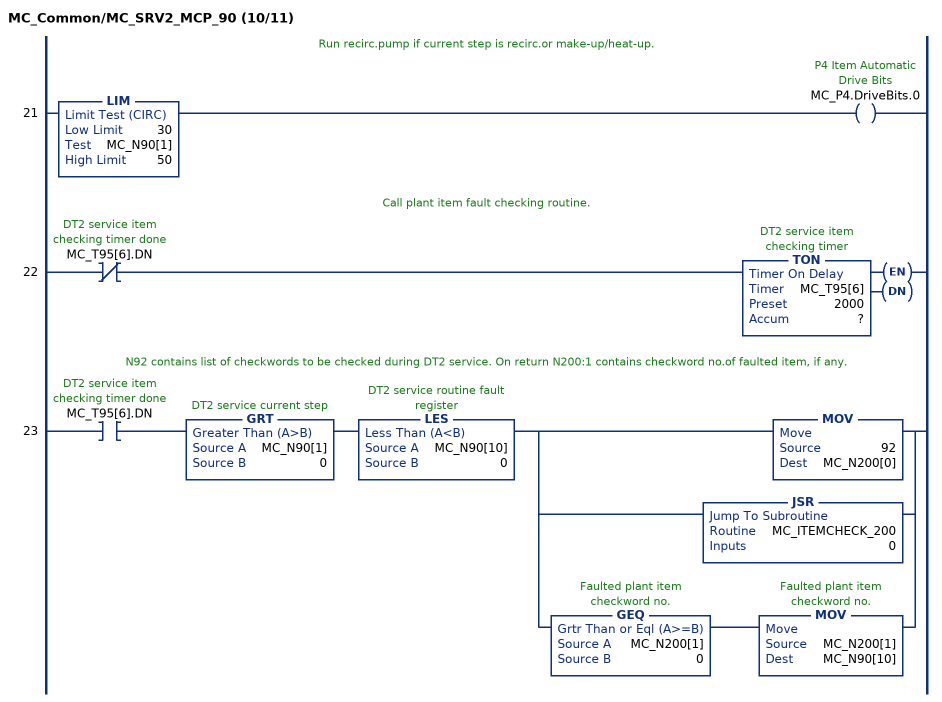
   // Run recirc.pump if current step is recirc.or make-up/heat-up.
   21: LIM(30,MC_N90[1],50)OTE(MC_P4.DriveBits.0);
   // Call plant item fault checking routine.
   22: XIO(MC_T95[6].DN)TON(MC_T95[6],?,?);
   // N92 contains list of checkwords to be checked during DT2 service. On return N200:1 contains checkword no.of faulted item, if any.
   23: XIC(MC_T95[6].DN)GRT(MC_N90[1],0)LES(MC_N90[10],0)[MOV(92,MC_N200[0]) ,JSR(MC_ITEMCHECK_200,0) ,GEQ(MC_N200[1],0) MOV(MC_N200[1],MC_N90[10]) ];
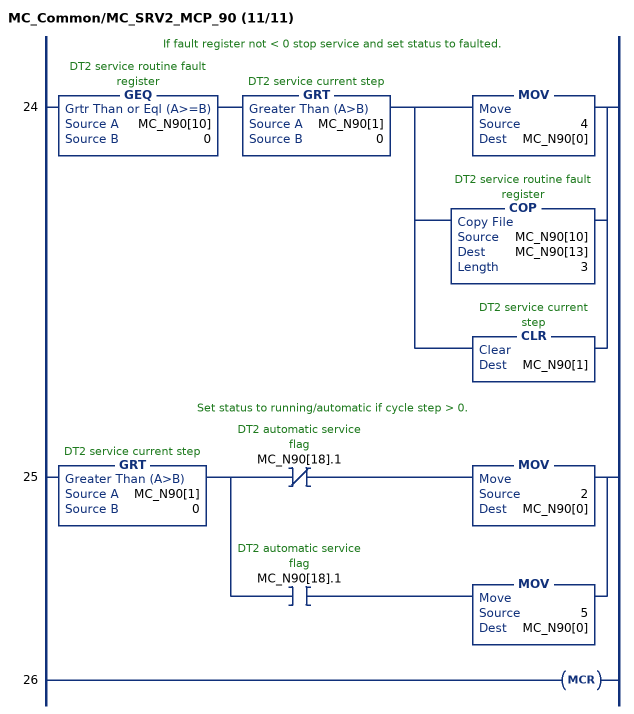
   // If fault register not < 0 stop service and set status to faulted.
   24: GEQ(MC_N90[10],0)GRT(MC_N90[1],0)[MOV(4,MC_N90[0]) ,COP(MC_N90[10],MC_N90[13],3) ,CLR(MC_N90[1]) ];
   // Set status to running/automatic if cycle step > 0.
   25: GRT(MC_N90[1],0)[XIO(MC_N90[18].1) MOV(2,MC_N90[0]) ,XIC(MC_N90[18].1) MOV(5,MC_N90[0]) ];
   26: MCR();
END_ROUTINE

ROUTINE MC_Valves   (* ladder *)
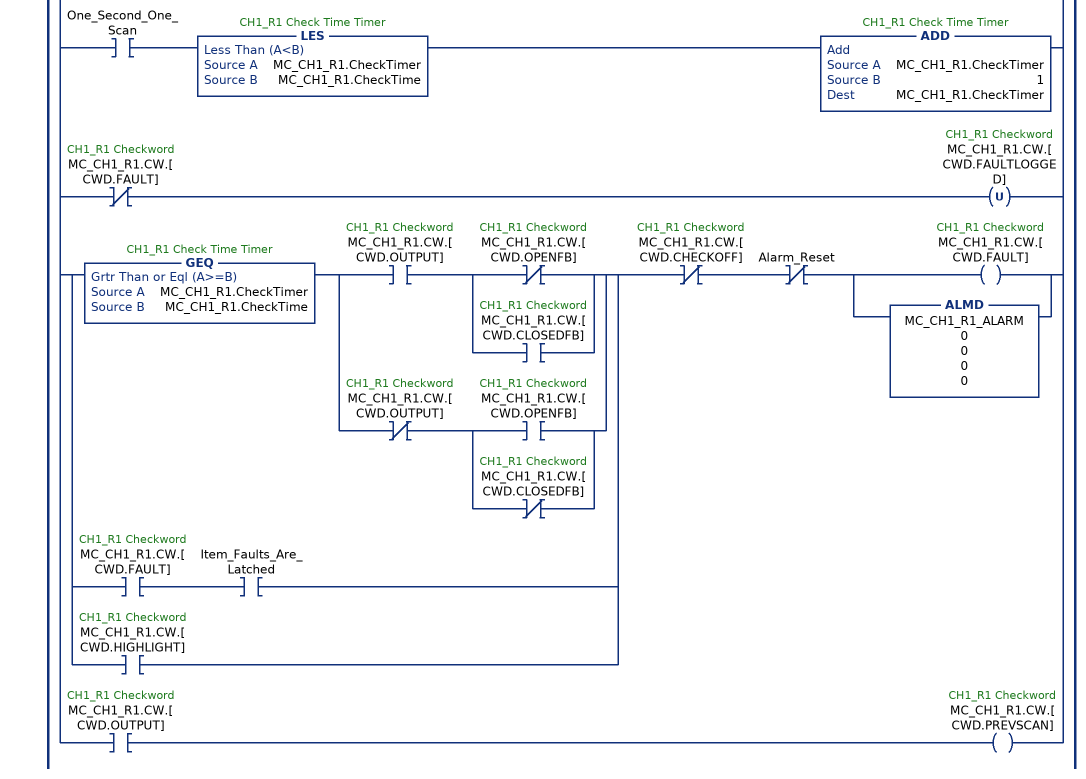
   0: [NEQ(MC_CH1_R1.DriveBits,0) OTE(MC_CH1_R1.CW.[CWD.AUTODRV]) ,[XIC(MC_CH1_R1.CW.[CWD.AUTODRV]) XIO(MC_CH1_R1.CW.[CWD.MANUAL]) ,XIC(MC_CH1_R1.CW.[CWD.MANDRV]) XIC(MC_CH1_R1.CW.[CWD.MANUAL]) ] OTE(MC_CH1_R1.CW.[CWD.OUTPUT]) ,XIC(MC_CH1_R1.CW.[CWD.OUTPUT]) OTE(MC_CH1_R1_DR) ,XIC(S:FS) [OTU(MC_CH1_R1.CW.[CWD.MANUAL]) ,LEQ(MC_CH1_R1.CheckTime,0) MOV(Default_Check_Time,MC_CH1_R1.CheckTime) ] ,[[XIC(MC_CH1_R1_O) XIO(Item_Simulation_Flag) ,XIC(Item_Simulation_Flag) XIC(MC_CH1_R1.CW.[CWD.OUTPUT]) XIO(MC_CH1_R1.CW.[CWD.SIMFAIL]) ] OTE(MC_CH1_R1.CW.[CWD.OPENFB]) ,[XIC(MC_CH1_R1_C) XIO(Item_Simulation_Flag) ,XIC(Item_Simulation_Flag) XIO(MC_CH1_R1.CW.[CWD.OUTPUT]) XIO(MC_CH1_R1.CW.[CWD.SIMFAIL]) ] OTE(MC_CH1_R1.CW.[CWD.CLOSEDFB]) ] ,[XIC(MC_CH1_R1.CW.[CWD.OUTPUT]) XIO(MC_CH1_R1.CW.[CWD.PREVSCAN]) ,XIO(MC_CH1_R1.CW.[CWD.OUTPUT]) XIC(MC_CH1_R1.CW.[CWD.PREVSCAN]) ] CLR(MC_CH1_R1.CheckTimer) ,XIC(One_Second_One_Scan) LES(MC_CH1_R1.CheckTimer,MC_CH1_R1.CheckTime) ADD(MC_CH1_R1.CheckTimer,1,MC_CH1_R1.CheckTimer) ,XIO(MC_CH1_R1.CW.[CWD.FAULT]) OTU(MC_CH1_R1.CW.[CWD.FAULTLOGGED]) ,[GEQ(MC_CH1_R1.CheckTimer,MC_CH1_R1.CheckTime) [XIC(MC_CH1_R1.CW.[CWD.OUTPUT]) [XIO(MC_CH1_R1.CW.[CWD.OPENFB]) ,XIC(MC_CH1_R1.CW.[CWD.CLOSEDFB]) ] ,XIO(MC_CH1_R1.CW.[CWD.OUTPUT]) [XIC(MC_CH1_R1.CW.[CWD.OPENFB]) ,XIO(MC_CH1_R1.CW.[CWD.CLOSEDFB]) ] ] ,XIC(MC_CH1_R1.CW.[CWD.FAULT]) XIC(Item_Faults_Are_Latched) ,XIC(MC_CH1_R1.CW.[CWD.HIGHLIGHT]) ] XIO(MC_CH1_R1.CW.[CWD.CHECKOFF]) XIO(Alarm_Reset) [OTE(MC_CH1_R1.CW.[CWD.FAULT]) ,ALMD(MC_CH1_R1_ALARM,0,0,0,0) ] ,XIC(MC_CH1_R1.CW.[CWD.OUTPUT]) OTE(MC_CH1_R1.CW.[CWD.PREVSCAN]) ];
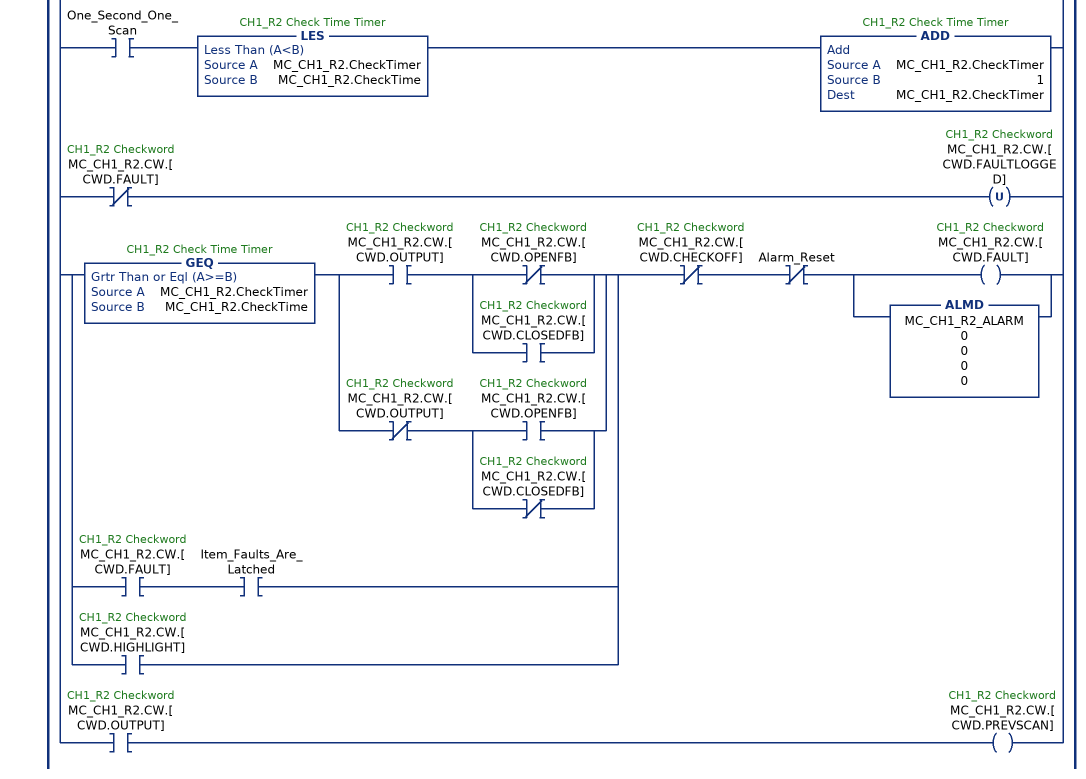
   1: [NEQ(MC_CH1_R2.DriveBits,0) OTE(MC_CH1_R2.CW.[CWD.AUTODRV]) ,[XIC(MC_CH1_R2.CW.[CWD.AUTODRV]) XIO(MC_CH1_R2.CW.[CWD.MANUAL]) ,XIC(MC_CH1_R2.CW.[CWD.MANDRV]) XIC(MC_CH1_R2.CW.[CWD.MANUAL]) ] OTE(MC_CH1_R2.CW.[CWD.OUTPUT]) ,XIC(MC_CH1_R2.CW.[CWD.OUTPUT]) OTE(MC_CH1_R2_DR) ,XIC(S:FS) [OTU(MC_CH1_R2.CW.[CWD.MANUAL]) ,LEQ(MC_CH1_R2.CheckTime,0) MOV(Default_Check_Time,MC_CH1_R2.CheckTime) ] ,[[XIC(MC_CH1_R2_O) XIO(Item_Simulation_Flag) ,XIC(Item_Simulation_Flag) XIC(MC_CH1_R2.CW.[CWD.OUTPUT]) XIO(MC_CH1_R2.CW.[CWD.SIMFAIL]) ] OTE(MC_CH1_R2.CW.[CWD.OPENFB]) ,[XIC(MC_CH1_R2_C) XIO(Item_Simulation_Flag) ,XIC(Item_Simulation_Flag) XIO(MC_CH1_R2.CW.[CWD.OUTPUT]) XIO(MC_CH1_R2.CW.[CWD.SIMFAIL]) ] OTE(MC_CH1_R2.CW.[CWD.CLOSEDFB]) ] ,[XIC(MC_CH1_R2.CW.[CWD.OUTPUT]) XIO(MC_CH1_R2.CW.[CWD.PREVSCAN]) ,XIO(MC_CH1_R2.CW.[CWD.OUTPUT]) XIC(MC_CH1_R2.CW.[CWD.PREVSCAN]) ] CLR(MC_CH1_R2.CheckTimer) ,XIC(One_Second_One_Scan) LES(MC_CH1_R2.CheckTimer,MC_CH1_R2.CheckTime) ADD(MC_CH1_R2.CheckTimer,1,MC_CH1_R2.CheckTimer) ,XIO(MC_CH1_R2.CW.[CWD.FAULT]) OTU(MC_CH1_R2.CW.[CWD.FAULTLOGGED]) ,[GEQ(MC_CH1_R2.CheckTimer,MC_CH1_R2.CheckTime) [XIC(MC_CH1_R2.CW.[CWD.OUTPUT]) [XIO(MC_CH1_R2.CW.[CWD.OPENFB]) ,XIC(MC_CH1_R2.CW.[CWD.CLOSEDFB]) ] ,XIO(MC_CH1_R2.CW.[CWD.OUTPUT]) [XIC(MC_CH1_R2.CW.[CWD.OPENFB]) ,XIO(MC_CH1_R2.CW.[CWD.CLOSEDFB]) ] ] ,XIC(MC_CH1_R2.CW.[CWD.FAULT]) XIC(Item_Faults_Are_Latched) ,XIC(MC_CH1_R2.CW.[CWD.HIGHLIGHT]) ] XIO(MC_CH1_R2.CW.[CWD.CHECKOFF]) XIO(Alarm_Reset) [OTE(MC_CH1_R2.CW.[CWD.FAULT]) ,ALMD(MC_CH1_R2_ALARM,0,0,0,0) ] ,XIC(MC_CH1_R2.CW.[CWD.OUTPUT]) OTE(MC_CH1_R2.CW.[CWD.PREVSCAN]) ];
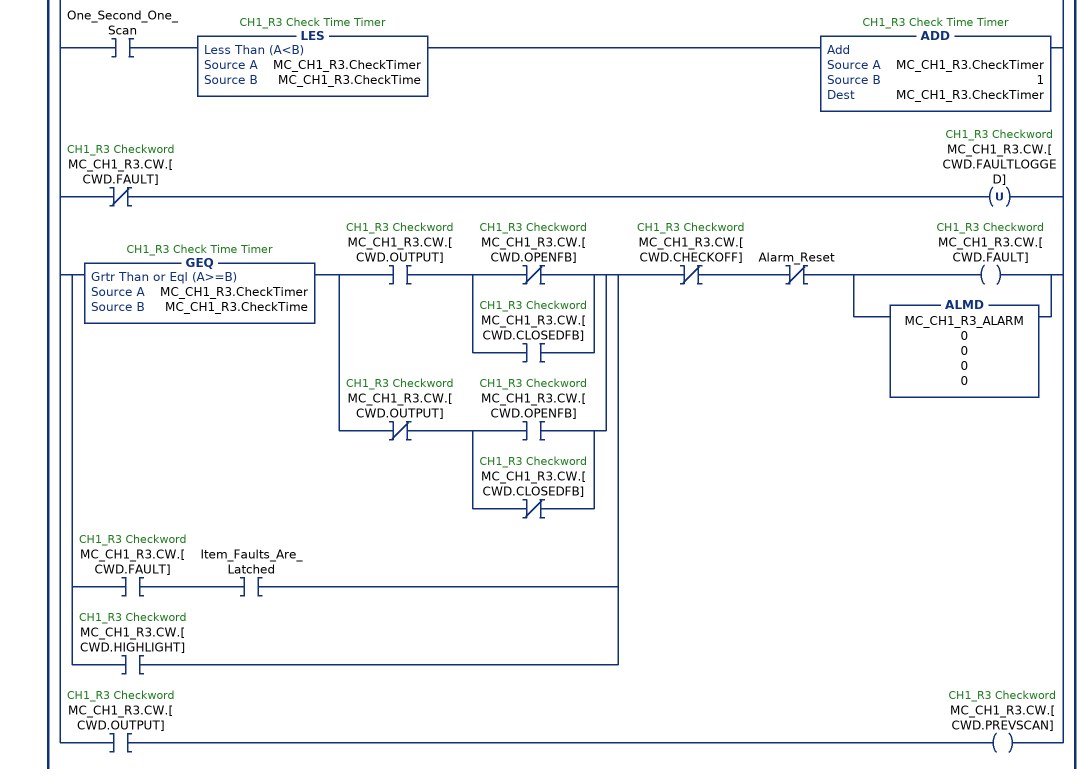
   2: [NEQ(MC_CH1_R3.DriveBits,0) OTE(MC_CH1_R3.CW.[CWD.AUTODRV]) ,[XIC(MC_CH1_R3.CW.[CWD.AUTODRV]) XIO(MC_CH1_R3.CW.[CWD.MANUAL]) ,XIC(MC_CH1_R3.CW.[CWD.MANDRV]) XIC(MC_CH1_R3.CW.[CWD.MANUAL]) ] OTE(MC_CH1_R3.CW.[CWD.OUTPUT]) ,XIC(MC_CH1_R3.CW.[CWD.OUTPUT]) OTE(MC_CH1_R3_DR) ,XIC(S:FS) [OTU(MC_CH1_R3.CW.[CWD.MANUAL]) ,LEQ(MC_CH1_R3.CheckTime,0) MOV(Default_Check_Time,MC_CH1_R3.CheckTime) ] ,[[XIC(MC_CH1_R3_O) XIO(Item_Simulation_Flag) ,XIC(Item_Simulation_Flag) XIC(MC_CH1_R3.CW.[CWD.OUTPUT]) XIO(MC_CH1_R3.CW.[CWD.SIMFAIL]) ] OTE(MC_CH1_R3.CW.[CWD.OPENFB]) ,[XIC(MC_CH1_R3_C) XIO(Item_Simulation_Flag) ,XIC(Item_Simulation_Flag) XIO(MC_CH1_R3.CW.[CWD.OUTPUT]) XIO(MC_CH1_R3.CW.[CWD.SIMFAIL]) ] OTE(MC_CH1_R3.CW.[CWD.CLOSEDFB]) ] ,[XIC(MC_CH1_R3.CW.[CWD.OUTPUT]) XIO(MC_CH1_R3.CW.[CWD.PREVSCAN]) ,XIO(MC_CH1_R3.CW.[CWD.OUTPUT]) XIC(MC_CH1_R3.CW.[CWD.PREVSCAN]) ] CLR(MC_CH1_R3.CheckTimer) ,XIC(One_Second_One_Scan) LES(MC_CH1_R3.CheckTimer,MC_CH1_R3.CheckTime) ADD(MC_CH1_R3.CheckTimer,1,MC_CH1_R3.CheckTimer) ,XIO(MC_CH1_R3.CW.[CWD.FAULT]) OTU(MC_CH1_R3.CW.[CWD.FAULTLOGGED]) ,[GEQ(MC_CH1_R3.CheckTimer,MC_CH1_R3.CheckTime) [XIC(MC_CH1_R3.CW.[CWD.OUTPUT]) [XIO(MC_CH1_R3.CW.[CWD.OPENFB]) ,XIC(MC_CH1_R3.CW.[CWD.CLOSEDFB]) ] ,XIO(MC_CH1_R3.CW.[CWD.OUTPUT]) [XIC(MC_CH1_R3.CW.[CWD.OPENFB]) ,XIO(MC_CH1_R3.CW.[CWD.CLOSEDFB]) ] ] ,XIC(MC_CH1_R3.CW.[CWD.FAULT]) XIC(Item_Faults_Are_Latched) ,XIC(MC_CH1_R3.CW.[CWD.HIGHLIGHT]) ] XIO(MC_CH1_R3.CW.[CWD.CHECKOFF]) XIO(Alarm_Reset) [OTE(MC_CH1_R3.CW.[CWD.FAULT]) ,ALMD(MC_CH1_R3_ALARM,0,0,0,0) ] ,XIC(MC_CH1_R3.CW.[CWD.OUTPUT]) OTE(MC_CH1_R3.CW.[CWD.PREVSCAN]) ];
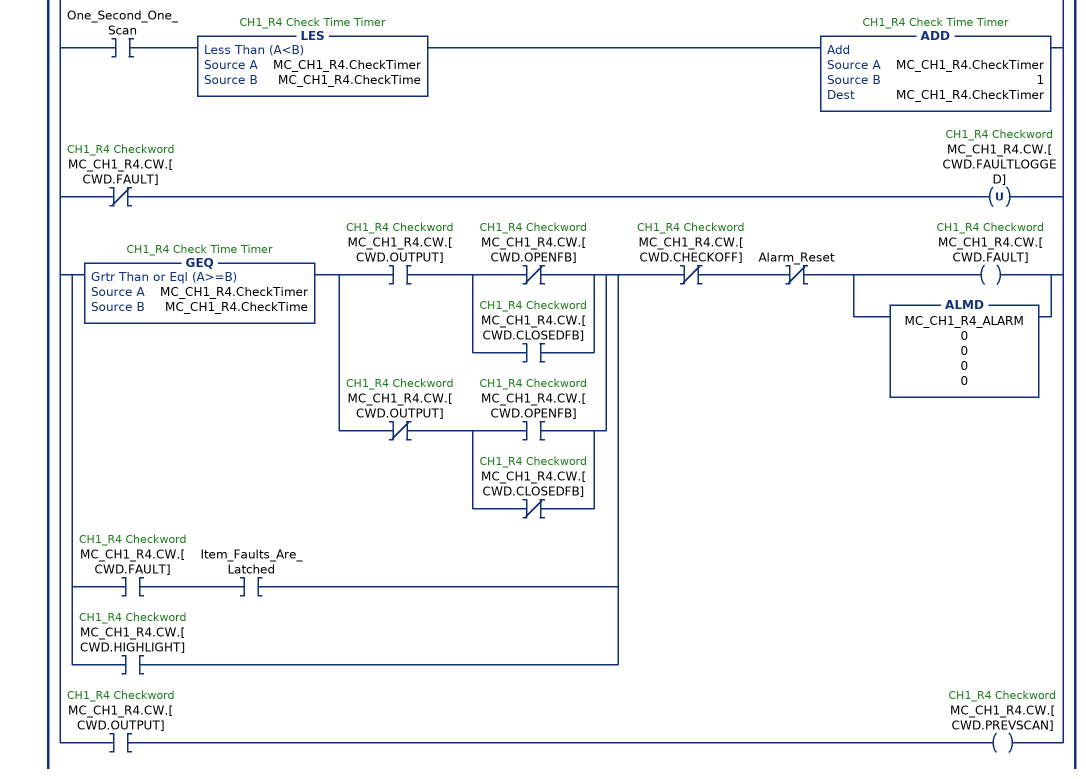
   3: [NEQ(MC_CH1_R4.DriveBits,0) OTE(MC_CH1_R4.CW.[CWD.AUTODRV]) ,[XIC(MC_CH1_R4.CW.[CWD.AUTODRV]) XIO(MC_CH1_R4.CW.[CWD.MANUAL]) ,XIC(MC_CH1_R4.CW.[CWD.MANDRV]) XIC(MC_CH1_R4.CW.[CWD.MANUAL]) ] OTE(MC_CH1_R4.CW.[CWD.OUTPUT]) ,XIC(MC_CH1_R4.CW.[CWD.OUTPUT]) OTE(MC_CH1_R4_DR) ,XIC(S:FS) [OTU(MC_CH1_R4.CW.[CWD.MANUAL]) ,LEQ(MC_CH1_R4.CheckTime,0) MOV(Default_Check_Time,MC_CH1_R4.CheckTime) ] ,[[XIC(MC_CH1_R4_O) XIO(Item_Simulation_Flag) ,XIC(Item_Simulation_Flag) XIC(MC_CH1_R4.CW.[CWD.OUTPUT]) XIO(MC_CH1_R4.CW.[CWD.SIMFAIL]) ] OTE(MC_CH1_R4.CW.[CWD.OPENFB]) ,[XIC(MC_CH1_R4_C) XIO(Item_Simulation_Flag) ,XIC(Item_Simulation_Flag) XIO(MC_CH1_R4.CW.[CWD.OUTPUT]) XIO(MC_CH1_R4.CW.[CWD.SIMFAIL]) ] OTE(MC_CH1_R4.CW.[CWD.CLOSEDFB]) ] ,[XIC(MC_CH1_R4.CW.[CWD.OUTPUT]) XIO(MC_CH1_R4.CW.[CWD.PREVSCAN]) ,XIO(MC_CH1_R4.CW.[CWD.OUTPUT]) XIC(MC_CH1_R4.CW.[CWD.PREVSCAN]) ] CLR(MC_CH1_R4.CheckTimer) ,XIC(One_Second_One_Scan) LES(MC_CH1_R4.CheckTimer,MC_CH1_R4.CheckTime) ADD(MC_CH1_R4.CheckTimer,1,MC_CH1_R4.CheckTimer) ,XIO(MC_CH1_R4.CW.[CWD.FAULT]) OTU(MC_CH1_R4.CW.[CWD.FAULTLOGGED]) ,[GEQ(MC_CH1_R4.CheckTimer,MC_CH1_R4.CheckTime) [XIC(MC_CH1_R4.CW.[CWD.OUTPUT]) [XIO(MC_CH1_R4.CW.[CWD.OPENFB]) ,XIC(MC_CH1_R4.CW.[CWD.CLOSEDFB]) ] ,XIO(MC_CH1_R4.CW.[CWD.OUTPUT]) [XIC(MC_CH1_R4.CW.[CWD.OPENFB]) ,XIO(MC_CH1_R4.CW.[CWD.CLOSEDFB]) ] ] ,XIC(MC_CH1_R4.CW.[CWD.FAULT]) XIC(Item_Faults_Are_Latched) ,XIC(MC_CH1_R4.CW.[CWD.HIGHLIGHT]) ] XIO(MC_CH1_R4.CW.[CWD.CHECKOFF]) XIO(Alarm_Reset) [OTE(MC_CH1_R4.CW.[CWD.FAULT]) ,ALMD(MC_CH1_R4_ALARM,0,0,0,0) ] ,XIC(MC_CH1_R4.CW.[CWD.OUTPUT]) OTE(MC_CH1_R4.CW.[CWD.PREVSCAN]) ];
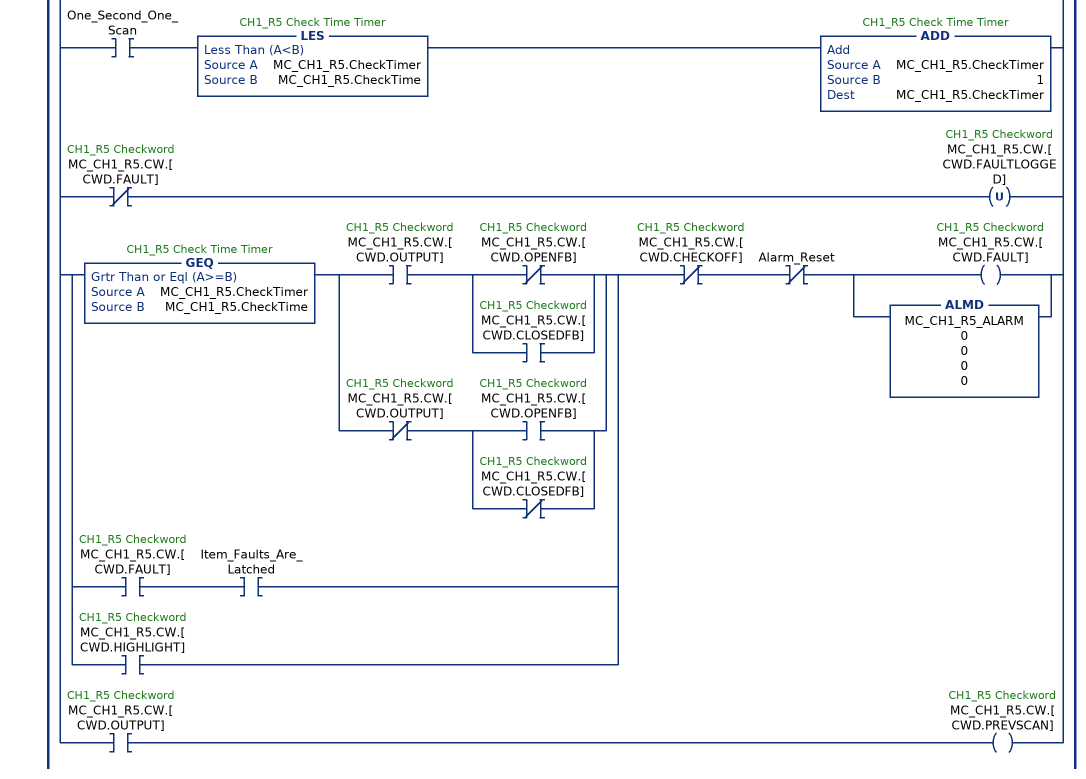
   4: [NEQ(MC_CH1_R5.DriveBits,0) OTE(MC_CH1_R5.CW.[CWD.AUTODRV]) ,[XIC(MC_CH1_R5.CW.[CWD.AUTODRV]) XIO(MC_CH1_R5.CW.[CWD.MANUAL]) ,XIC(MC_CH1_R5.CW.[CWD.MANDRV]) XIC(MC_CH1_R5.CW.[CWD.MANUAL]) ] OTE(MC_CH1_R5.CW.[CWD.OUTPUT]) ,XIC(MC_CH1_R5.CW.[CWD.OUTPUT]) OTE(MC_CH1_R5_DR) ,XIC(S:FS) [OTU(MC_CH1_R5.CW.[CWD.MANUAL]) ,LEQ(MC_CH1_R5.CheckTime,0) MOV(Default_Check_Time,MC_CH1_R5.CheckTime) ] ,[[XIC(MC_CH1_R5_O) XIO(Item_Simulation_Flag) ,XIC(Item_Simulation_Flag) XIC(MC_CH1_R5.CW.[CWD.OUTPUT]) XIO(MC_CH1_R5.CW.[CWD.SIMFAIL]) ] OTE(MC_CH1_R5.CW.[CWD.OPENFB]) ,[XIC(MC_CH1_R5_C) XIO(Item_Simulation_Flag) ,XIC(Item_Simulation_Flag) XIO(MC_CH1_R5.CW.[CWD.OUTPUT]) XIO(MC_CH1_R5.CW.[CWD.SIMFAIL]) ] OTE(MC_CH1_R5.CW.[CWD.CLOSEDFB]) ] ,[XIC(MC_CH1_R5.CW.[CWD.OUTPUT]) XIO(MC_CH1_R5.CW.[CWD.PREVSCAN]) ,XIO(MC_CH1_R5.CW.[CWD.OUTPUT]) XIC(MC_CH1_R5.CW.[CWD.PREVSCAN]) ] CLR(MC_CH1_R5.CheckTimer) ,XIC(One_Second_One_Scan) LES(MC_CH1_R5.CheckTimer,MC_CH1_R5.CheckTime) ADD(MC_CH1_R5.CheckTimer,1,MC_CH1_R5.CheckTimer) ,XIO(MC_CH1_R5.CW.[CWD.FAULT]) OTU(MC_CH1_R5.CW.[CWD.FAULTLOGGED]) ,[GEQ(MC_CH1_R5.CheckTimer,MC_CH1_R5.CheckTime) [XIC(MC_CH1_R5.CW.[CWD.OUTPUT]) [XIO(MC_CH1_R5.CW.[CWD.OPENFB]) ,XIC(MC_CH1_R5.CW.[CWD.CLOSEDFB]) ] ,XIO(MC_CH1_R5.CW.[CWD.OUTPUT]) [XIC(MC_CH1_R5.CW.[CWD.OPENFB]) ,XIO(MC_CH1_R5.CW.[CWD.CLOSEDFB]) ] ] ,XIC(MC_CH1_R5.CW.[CWD.FAULT]) XIC(Item_Faults_Are_Latched) ,XIC(MC_CH1_R5.CW.[CWD.HIGHLIGHT]) ] XIO(MC_CH1_R5.CW.[CWD.CHECKOFF]) XIO(Alarm_Reset) [OTE(MC_CH1_R5.CW.[CWD.FAULT]) ,ALMD(MC_CH1_R5_ALARM,0,0,0,0) ] ,XIC(MC_CH1_R5.CW.[CWD.OUTPUT]) OTE(MC_CH1_R5.CW.[CWD.PREVSCAN]) ];
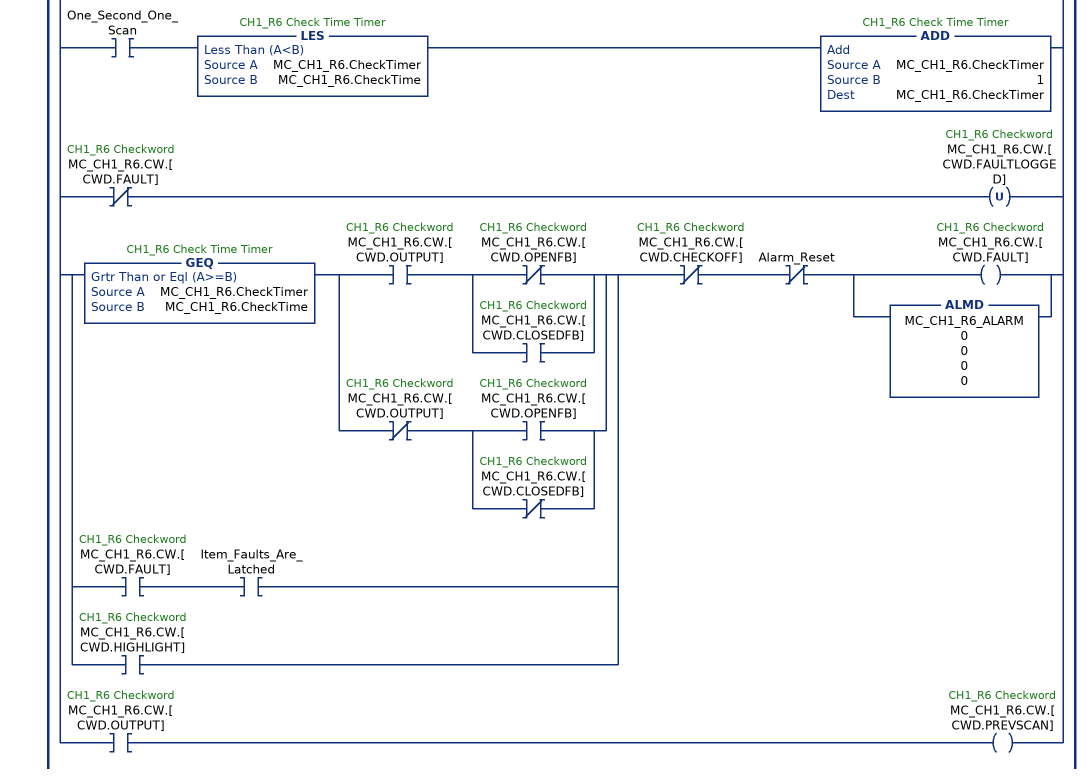
   5: [NEQ(MC_CH1_R6.DriveBits,0) OTE(MC_CH1_R6.CW.[CWD.AUTODRV]) ,[XIC(MC_CH1_R6.CW.[CWD.AUTODRV]) XIO(MC_CH1_R6.CW.[CWD.MANUAL]) ,XIC(MC_CH1_R6.CW.[CWD.MANDRV]) XIC(MC_CH1_R6.CW.[CWD.MANUAL]) ] OTE(MC_CH1_R6.CW.[CWD.OUTPUT]) ,XIC(MC_CH1_R6.CW.[CWD.OUTPUT]) OTE(MC_CH1_R6_DR) ,XIC(S:FS) [OTU(MC_CH1_R6.CW.[CWD.MANUAL]) ,LEQ(MC_CH1_R6.CheckTime,0) MOV(Default_Check_Time,MC_CH1_R6.CheckTime) ] ,[[XIC(MC_CH1_R6_O) XIO(Item_Simulation_Flag) ,XIC(Item_Simulation_Flag) XIC(MC_CH1_R6.CW.[CWD.OUTPUT]) XIO(MC_CH1_R6.CW.[CWD.SIMFAIL]) ] OTE(MC_CH1_R6.CW.[CWD.OPENFB]) ,[XIC(MC_CH1_R6_C) XIO(Item_Simulation_Flag) ,XIC(Item_Simulation_Flag) XIO(MC_CH1_R6.CW.[CWD.OUTPUT]) XIO(MC_CH1_R6.CW.[CWD.SIMFAIL]) ] OTE(MC_CH1_R6.CW.[CWD.CLOSEDFB]) ] ,[XIC(MC_CH1_R6.CW.[CWD.OUTPUT]) XIO(MC_CH1_R6.CW.[CWD.PREVSCAN]) ,XIO(MC_CH1_R6.CW.[CWD.OUTPUT]) XIC(MC_CH1_R6.CW.[CWD.PREVSCAN]) ] CLR(MC_CH1_R6.CheckTimer) ,XIC(One_Second_One_Scan) LES(MC_CH1_R6.CheckTimer,MC_CH1_R6.CheckTime) ADD(MC_CH1_R6.CheckTimer,1,MC_CH1_R6.CheckTimer) ,XIO(MC_CH1_R6.CW.[CWD.FAULT]) OTU(MC_CH1_R6.CW.[CWD.FAULTLOGGED]) ,[GEQ(MC_CH1_R6.CheckTimer,MC_CH1_R6.CheckTime) [XIC(MC_CH1_R6.CW.[CWD.OUTPUT]) [XIO(MC_CH1_R6.CW.[CWD.OPENFB]) ,XIC(MC_CH1_R6.CW.[CWD.CLOSEDFB]) ] ,XIO(MC_CH1_R6.CW.[CWD.OUTPUT]) [XIC(MC_CH1_R6.CW.[CWD.OPENFB]) ,XIO(MC_CH1_R6.CW.[CWD.CLOSEDFB]) ] ] ,XIC(MC_CH1_R6.CW.[CWD.FAULT]) XIC(Item_Faults_Are_Latched) ,XIC(MC_CH1_R6.CW.[CWD.HIGHLIGHT]) ] XIO(MC_CH1_R6.CW.[CWD.CHECKOFF]) XIO(Alarm_Reset) [OTE(MC_CH1_R6.CW.[CWD.FAULT]) ,ALMD(MC_CH1_R6_ALARM,0,0,0,0) ] ,XIC(MC_CH1_R6.CW.[CWD.OUTPUT]) OTE(MC_CH1_R6.CW.[CWD.PREVSCAN]) ];
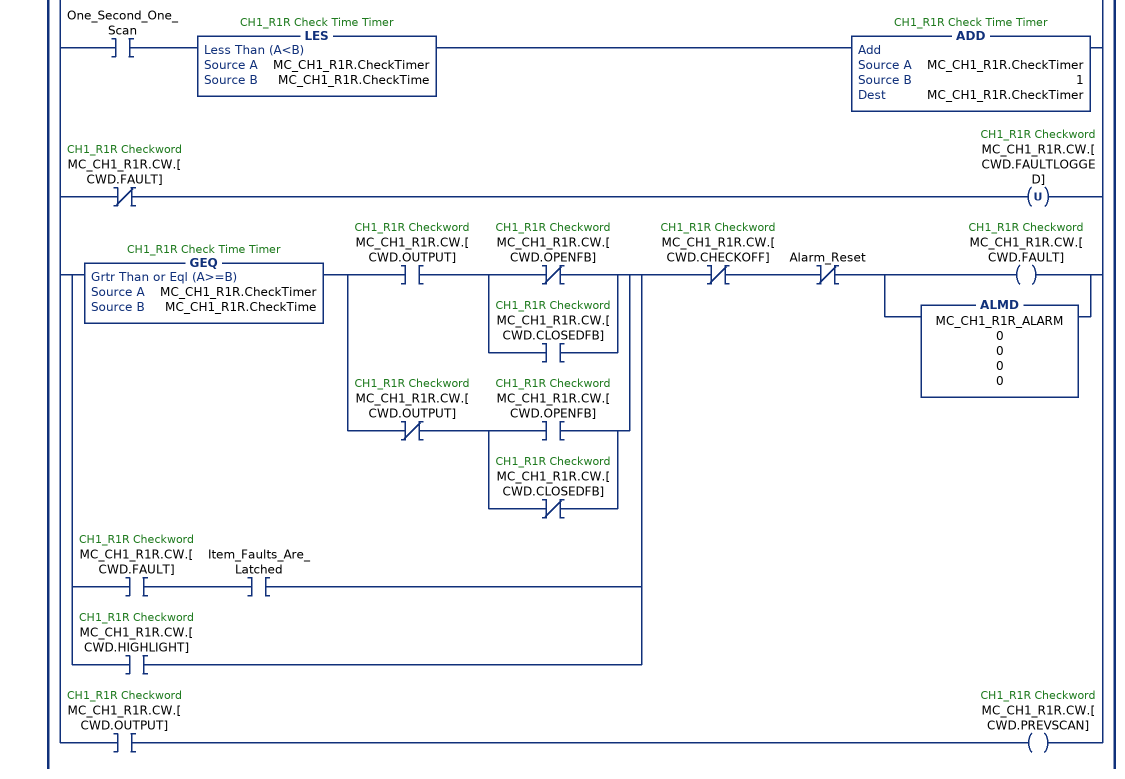
   6: [NEQ(MC_CH1_R1R.DriveBits,0) OTE(MC_CH1_R1R.CW.[CWD.AUTODRV]) ,[XIC(MC_CH1_R1R.CW.[CWD.AUTODRV]) XIO(MC_CH1_R1R.CW.[CWD.MANUAL]) ,XIC(MC_CH1_R1R.CW.[CWD.MANDRV]) XIC(MC_CH1_R1R.CW.[CWD.MANUAL]) ] OTE(MC_CH1_R1R.CW.[CWD.OUTPUT]) ,XIC(MC_CH1_R1R.CW.[CWD.OUTPUT]) OTE(MC_CH1_R1R_DR) ,XIC(S:FS) [OTU(MC_CH1_R1R.CW.[CWD.MANUAL]) ,LEQ(MC_CH1_R1R.CheckTime,0) MOV(Default_Check_Time,MC_CH1_R1R.CheckTime) ] ,[[XIC(MC_CH1_R1R_O) XIO(Item_Simulation_Flag) ,XIC(Item_Simulation_Flag) XIC(MC_CH1_R1R.CW.[CWD.OUTPUT]) XIO(MC_CH1_R1R.CW.[CWD.SIMFAIL]) ] OTE(MC_CH1_R1R.CW.[CWD.OPENFB]) ,[XIC(MC_CH1_R1R_C) XIO(Item_Simulation_Flag) ,XIC(Item_Simulation_Flag) XIO(MC_CH1_R1R.CW.[CWD.OUTPUT]) XIO(MC_CH1_R1R.CW.[CWD.SIMFAIL]) ] OTE(MC_CH1_R1R.CW.[CWD.CLOSEDFB]) ] ,[XIC(MC_CH1_R1R.CW.[CWD.OUTPUT]) XIO(MC_CH1_R1R.CW.[CWD.PREVSCAN]) ,XIO(MC_CH1_R1R.CW.[CWD.OUTPUT]) XIC(MC_CH1_R1R.CW.[CWD.PREVSCAN]) ] CLR(MC_CH1_R1R.CheckTimer) ,XIC(One_Second_One_Scan) LES(MC_CH1_R1R.CheckTimer,MC_CH1_R1R.CheckTime) ADD(MC_CH1_R1R.CheckTimer,1,MC_CH1_R1R.CheckTimer) ,XIO(MC_CH1_R1R.CW.[CWD.FAULT]) OTU(MC_CH1_R1R.CW.[CWD.FAULTLOGGED]) ,[GEQ(MC_CH1_R1R.CheckTimer,MC_CH1_R1R.CheckTime) [XIC(MC_CH1_R1R.CW.[CWD.OUTPUT]) [XIO(MC_CH1_R1R.CW.[CWD.OPENFB]) ,XIC(MC_CH1_R1R.CW.[CWD.CLOSEDFB]) ] ,XIO(MC_CH1_R1R.CW.[CWD.OUTPUT]) [XIC(MC_CH1_R1R.CW.[CWD.OPENFB]) ,XIO(MC_CH1_R1R.CW.[CWD.CLOSEDFB]) ] ] ,XIC(MC_CH1_R1R.CW.[CWD.FAULT]) XIC(Item_Faults_Are_Latched) ,XIC(MC_CH1_R1R.CW.[CWD.HIGHLIGHT]) ] XIO(MC_CH1_R1R.CW.[CWD.CHECKOFF]) XIO(Alarm_Reset) [OTE(MC_CH1_R1R.CW.[CWD.FAULT]) ,ALMD(MC_CH1_R1R_ALARM,0,0,0,0) ] ,XIC(MC_CH1_R1R.CW.[CWD.OUTPUT]) OTE(MC_CH1_R1R.CW.[CWD.PREVSCAN]) ];
